DATA_BLOCK "DB_Z256_Scada"   // DB2010
{ S7_Optimized_Access := 'FALSE' }
VERSION : 0.1
   VAR
      tAlm : Struct   // HMI Alarms
         tE : Struct
            x0 : Bool;   // KE.Main emergency on
            x1 : Bool;   // KE1.Local emergency on
            x2 : Bool;   // Cabinet.Emergency localization
            x3 : Bool;   // SB1.Emergency localization
            x4 : Bool;   // SB2.Emergency localization
            x5 : Bool;
            x6 : Bool;
            x7 : Bool;
            x8 : Bool;
            x9 : Bool;
            x10 : Bool;
            x11 : Bool;
            x12 : Bool;
            x13 : Bool;
            x14 : Bool;
            x15 : Bool;
            x16 : Bool;
            x17 : Bool;
            x18 : Bool;
            x19 : Bool;
            x20 : Bool;
            x21 : Bool;
            x22 : Bool;
            x23 : Bool;
            x24 : Bool;
            x25 : Bool;
            x26 : Bool;
            x27 : Bool;
            x28 : Bool;
            x29 : Bool;
            x30 : Bool;
            x31 : Bool;
         END_STRUCT;
         tS : Struct
            tS0 : Struct
               x0 : Bool;   // xB18-3L+.PowerSupplyInputControlCabinetON
               x1 : Bool;   // xB18-7L+.InputInstallationPowerSupplyON"
               x2 : Bool;   // xB11QF1/1D/QF2.Anomaly power supplies 120V
               x3 : Bool;   // xB115KM1/2.AuxiliaryPowerSupplySetIn / xB18QF2.Power supply 24V logic
               x4 : Bool;   // xB410AP1.SafetyOnPanel1" / xB18QF3.Power supply 24V logic
               x5 : Bool;   // xB410AP1.SafetyOnPanel2" / xB20QF2.Power supply 24V logic
               x6 : Bool;   // xB20QF3.Power supply 24V logic
               x7 : Bool;   // xB21QF1.Power supply 24V logic
               x8 : Bool;   // xB140QF2.ProtectionPowerSupplyMotorsYcut" / xB41QF1.ProtectionPowerSupplyMotorsYcut 1-4
               x9 : Bool;   // xB41QF2.Protection power supply motors longitudinal cutting / xB41QF2.Protection power supply 36V motors longitudinal cutting 1-4
               x10 : Bool;   // xB42QF1.Protection power supply 36V / xB42QF1.ProtectionPowerSupplyMotorsYcut 5-8
               x11 : Bool;   // xB42QF2.Protection power supply motors longitudinal cutting / xB42QF2.Protection power supply 36V motors longitudinal cutting 5-8
               x12 : Bool;
               x13 : Bool;
               x14 : Bool;
               x15 : Bool;
               x16 : Bool;   // PLCA.Timeout receiving consumed message
               x17 : Bool;   // PLCB.Timeout receiving consumed message
               x18 : Bool;   // PLCA.Mission packet lost
               x19 : Bool;   // PLCB.Mission packet lost
               x20 : Bool;   // PLCA.Syncro packet lost
               x21 : Bool;   // PLCB.Syncro packet lost
               x22 : Bool;   // Syncro.YCut meter gap outside the limits
               x23 : Bool;   // Syncro.Main line meter gap outside the limits
               x24 : Bool;   // Syncro.Timeout receiving meter signal from main line
               x25 : Bool;   // Syncro.Timeout receiving syncro value from mainline
               x26 : Bool;   // Syncro.Unexpected syncro pulse
               x27 : Bool;   // Syncro.Unexpected syncro message
               x28 : Bool;   // Syncro.Machine not syncronized
               x29 : Bool;
               x30 : Bool;
               x31 : Bool;
            END_STRUCT;
            tS1 : Struct
               x0 : Bool;
               x1 : Bool;   // Syncro.YCut meter gap outside the limits
               x2 : Bool;
               x3 : Bool;
               x4 : Bool;
               x5 : Bool;
               x6 : Bool;
               x7 : Bool;
               x8 : Bool;   // xB21QF1.Power supply 24V logic
               x9 : Bool;
               x10 : Bool;   // Syncro.Main line meter gap outside the limits
               x11 : Bool;
               x12 : Bool;
               x13 : Bool;
               x14 : Bool;
               x15 : Bool;
               x16 : Bool;
               x17 : Bool;
               x18 : Bool;
               x19 : Bool;
               x20 : Bool;
               x21 : Bool;
               x22 : Bool;
               x23 : Bool;
               x24 : Bool;
               x25 : Bool;
               x26 : Bool;
               x27 : Bool;
               x28 : Bool;
               x29 : Bool;
               x30 : Bool;
               x31 : Bool;
            END_STRUCT;
            tS2 : Struct
               x0 : Bool;
               x1 : Bool;   // Syncro.YCut meter gap outside the limits
               x2 : Bool;
               x3 : Bool;
               x4 : Bool;
               x5 : Bool;
               x6 : Bool;
               x7 : Bool;
               x8 : Bool;   // xB21QF1.Power supply 24V logic
               x9 : Bool;
               x10 : Bool;   // Syncro.Main line meter gap outside the limits
               x11 : Bool;
               x12 : Bool;
               x13 : Bool;
               x14 : Bool;
               x15 : Bool;
               x16 : Bool;
               x17 : Bool;
               x18 : Bool;
               x19 : Bool;
               x20 : Bool;
               x21 : Bool;
               x22 : Bool;
               x23 : Bool;
               x24 : Bool;
               x25 : Bool;
               x26 : Bool;
               x27 : Bool;
               x28 : Bool;
               x29 : Bool;
               x30 : Bool;
               x31 : Bool;
            END_STRUCT;
            tS3 : Struct
               x0 : Bool;
               x1 : Bool;   // Syncro.YCut meter gap outside the limits
               x2 : Bool;
               x3 : Bool;
               x4 : Bool;
               x5 : Bool;
               x6 : Bool;
               x7 : Bool;
               x8 : Bool;   // xB21QF1.Power supply 24V logic
               x9 : Bool;
               x10 : Bool;   // Syncro.Main line meter gap outside the limits
               x11 : Bool;
               x12 : Bool;
               x13 : Bool;
               x14 : Bool;
               x15 : Bool;
               x16 : Bool;
               x17 : Bool;
               x18 : Bool;
               x19 : Bool;
               x20 : Bool;
               x21 : Bool;
               x22 : Bool;
               x23 : Bool;
               x24 : Bool;
               x25 : Bool;
               x26 : Bool;
               x27 : Bool;
               x28 : Bool;
               x29 : Bool;
               x30 : Bool;
               x31 : Bool;
            END_STRUCT;
         END_STRUCT;
         tF : Struct
            x0 : Bool;
            x1 : Bool;
            x2 : Bool;
            x3 : Bool;
            x4 : Bool;
            x5 : Bool;
            x6 : Bool;
            x7 : Bool;
            x8 : Bool;
            x9 : Bool;
            x10 : Bool;
            x11 : Bool;
            x12 : Bool;
            x13 : Bool;
            x14 : Bool;
            x15 : Bool;
            x16 : Bool;
            x17 : Bool;
            x18 : Bool;
            x19 : Bool;
            x20 : Bool;
            x21 : Bool;
            x22 : Bool;
            x23 : Bool;
            x24 : Bool;
            x25 : Bool;
            x26 : Bool;
            x27 : Bool;
            x28 : Bool;
            x29 : Bool;
            x30 : Bool;
            x31 : Bool;
         END_STRUCT;
         tW : Struct
            x0 : Bool;   // PLCA.Timeout receiving consumed message
            x1 : Bool;   // PLCB.Timeout receiving consumed message
            x2 : Bool;   // PLCA.Mission packet lost
            x3 : Bool;   // PLCB.Mission packet lost
            x4 : Bool;   // PLCA.Syncro packet lost
            x5 : Bool;   // PLCB.Syncro packet lost
            x6 : Bool;   // QF.Protection air conditioners
            x7 : Bool;
            x8 : Bool;
            x9 : Bool;
            x10 : Bool;
            x11 : Bool;
            x12 : Bool;
            x13 : Bool;
            x14 : Bool;
            x15 : Bool;
            x16 : Bool;
            x17 : Bool;
            x18 : Bool;
            x19 : Bool;
            x20 : Bool;
            x21 : Bool;
            x22 : Bool;
            x23 : Bool;
            x24 : Bool;
            x25 : Bool;
            x26 : Bool;
            x27 : Bool;
            x28 : Bool;
            x29 : Bool;
            x30 : Bool;
            x31 : Bool;
         END_STRUCT;
      END_STRUCT;
      tHMR : Struct   // HMI Read
         xCalibrationsAllowed : Bool := FALSE;   // Calibration function allowed {x|x|x|x|O}
         xSpare1 : Bool;
         xSpare2 : Bool;
         xSpare3 : Bool;
         xSpare4 : Bool;
         xSpare5 : Bool;
         xSpare6 : Bool;
         xSpare7 : Bool;
         xSpare8 : Bool;
         xSpare9 : Bool;
         xSpare10 : Bool;
         xSpare11 : Bool;
         xSpare12 : Bool;
         xSpare13 : Bool;
         xSpare14 : Bool;
         xZoneAlarm : Bool := FALSE;   // Zone alarm {X|X|X|X|O}
         xSpare16 : Bool;
         xSpare17 : Bool;
         xSpare18 : Bool;
         xSpare19 : Bool;
         xSpare20 : Bool;
         xSpare21 : Bool;
         xSpare22 : Bool;
         xSpare23 : Bool;
         xSpare24 : Bool;
         xSpare25 : Bool;
         xSpare26 : Bool;
         xSpare27 : Bool;
         xSpare28 : Bool;
         xSpare29 : Bool;
         xSpare30 : Bool;
         xSpare31 : Bool;
         xSpare : Array[0..15] of Bool;
         iSpare0 : Int;
         iSpare1 : Int;
         iSpare2 : Int;
         iSpare3 : Int;
         iSpare4 : Int;
         iSpare5 : Int;
         iSpare6 : Int;
         iSpare7 : Int;
         iSpare8 : Int;
         iSpare9 : Int;
         iSpare10 : Int;
         iSpare11 : Int;
         iSpare12 : Int;
         iSpare13 : Int;
         iSpare14 : Int;
         iSpare15 : Int;
         iSpare16 : Int;
         dZoneMode : DInt := 4;   // Zone modality (1=Manual;4=Automatic;8=Manual request) {x|x|x|x|O}
         dZoneState : DInt := 1024;   // Zone status (1=CycleON 2=StopCyc 4=CycleReq 8=StopReq 1024=E-Stop) {X|X|X|X|O} / HMI Alarms
         dCabinetStatusMCC : DInt := 1;   // Cabinet status MCC1256B (1=OK;2=General power alarm;3=Local power alarm) {X|X|X|X|O} / HMI Write
         dProdModeRequest : DInt := 3;   // Production modality request (1=Out of Production 3= In production) {x|x|x|x|O}
         dProdModeActual : DInt := 3;   // Production modality actual (1=Out of production 3=In production 8=Out of production request 9=In production request) {x|x|x|x|O}
         dSpare5 : DInt;
         "rgdHeadsActualStatus[0]" : DInt := 3;   // Head #1 prod. status (1=Out of production 3=In production 8=Out of production request 9=In production request) {x|x|x|x|O}
         "rgdHeadsActualStatus[1]" : DInt := 3;   // Head #2 prod. status (1=Out of production 3=In production 8=Out of production request 9=In production request) {x|x|x|x|O}
         "rgdHeadsActualStatus[2]" : DInt := 3;   // Head #3 prod. status (1=Out of production 3=In production 8=Out of production request 9=In production request) {x|x|x|x|O}
         "rgdHeadsActualStatus[3]" : DInt := 3;   // Head #4 prod. status (1=Out of production 3=In production 8=Out of production request 9=In production request) {x|x|x|x|O}
         "rgdHeadsActualStatus[4]" : DInt;   // Head #5 prod. status (1=Out of production 3=In production 8=Out of production request 9=In production request) {x|x|x|x|O}
         "rgdHeadsActualStatus[5]" : DInt;   // Head #6 prod. status (1=Out of production 3=In production 8=Out of production request 9=In production request) {x|x|x|x|O}
         "rgdHeadsActualStatus[6]" : DInt;   // Head #7 prod. status (1=Out of production 3=In production 8=Out of production request 9=In production request) {x|x|x|x|O}
         "rgdHeadsActualStatus[7]" : DInt;   // Head #8 prod. status (1=Out of production 3=In production 8=Out of production request 9=In production request) {x|x|x|x|O}
         dSpare14 : DInt;
         dSpare15 : DInt;
         dSpare : Array[0..15] of DInt;
         rSpare0 : Real;
         rSpare1 : Real;
         rSpare2 : Real;
         rSpare3 : Real;
         rSpare4 : Real;
         rSpare5 : Real;
         rSpare6 : Real;
         rSpare7 : Real;
         rSpare8 : Real;
         tManCmd : Struct
            xSpare0 : Bool;
            xSpare1 : Bool;
            xSpare2 : Bool;
            xSpare3 : Bool;
            xSpare4 : Bool;
            xSpare5 : Bool;
            xSpare6 : Bool;
            xSpare7 : Bool;
            xSpare8 : Bool;
            xSpare9 : Bool;
            xSpare10 : Bool;
            xSpare11 : Bool;
            xSpare12 : Bool;
            xSpare13 : Bool;
            xSpare14 : Bool;
            xSpare15 : Bool;
            xSpare : Array[0..15] of Bool;
         END_STRUCT;
      END_STRUCT;
      tHMW : Struct   // HMI Write
         xAutoModeReq : Bool := FALSE;   // Automatic mode request {x|x|x|x|O}
         xManModeReq : Bool := FALSE;   // Manual mode request {x|x|x|x|O}
         xOutOfProdReq : Bool := FALSE;   // Bridge out of production request {x|x|x|x|O}
         xInProdReq : Bool := FALSE;   // Bridge in production request {x|x|x|x|O}
         xCutOnBreakEnabled : Bool := FALSE;   // Cut during glass break {x|x|x|x|O}
         xMotorsAndCardsInitialize : Bool := FALSE;   // Motors and cards initialize {x|x|x|x|M}
         xForceHeadsHoming : Bool := FALSE;   // Force the homing of the heads {x|x|x|x|M}
         xPositionCalibrationRequest : Bool := FALSE;   // Position calibration request {x|x|x|x|M}
         xBridgeOffsetCalibrationRequest : Bool := FALSE;   // Bridge offset calibration request {x|x|x|x|M}
         xSpare9 : Bool;
         xSpare10 : Bool;
         xSpare11 : Bool;
         xSpare12 : Bool;
         xSpare13 : Bool;
         xGeneralReset : Bool := FALSE;   // General reset {X|X|X|X|M}
         xFaultsReset : Bool := FALSE;   // Reset faults {X|X|X|X|O}
         xHeadEnabled_1 : Bool := TRUE;   // Head #1 enabled/disabled {x|x|x|x|O}
         xHeadEnabled_2 : Bool := TRUE;   // Head #2 enabled/disabled {x|x|x|x|O}
         xHeadEnabled_3 : Bool := TRUE;   // Head #3 enabled/disabled {x|x|x|x|O}
         xHeadEnabled_4 : Bool := TRUE;   // Head #4 enabled/disabled {x|x|x|x|O}
         xHeadEnabled_5 : Bool := TRUE;   // Head #5 enabled/disabled {x|x|x|x|O}
         xHeadEnabled_6 : Bool := TRUE;   // Head #6 enabled/disabled {x|x|x|x|O}
         xHeadEnabled_7 : Bool := TRUE;   // Head #7 enabled/disabled {x|x|x|x|O}
         xHeadEnabled_8 : Bool := TRUE;   // Head #8 enabled/disabled {x|x|x|x|O}
         xSpare24 : Bool;
         xSpare25 : Bool;
         xSpare26 : Bool;
         xSpare27 : Bool;
         xSpare28 : Bool;
         xSpare29 : Bool;
         xSpare30 : Bool;
         xSpare31 : Bool;
         xSpare : Array[0..15] of Bool;
         iSpare0 : Int;
         iSpare1 : Int;
         iSpare2 : Int;
         iSpare3 : Int;
         iSpare4 : Int;
         iSpare5 : Int;
         iSpare6 : Int;
         iSpare7 : Int;
         iSpare8 : Int;
         iSpare9 : Int;
         iSpare10 : Int;
         iSpare11 : Int;
         iSpare12 : Int;
         iSpare13 : Int;
         iSpare14 : Int;
         iSpare15 : Int;
         iSpare16 : Int;
         dNumberOfLites : DInt := 1;   // Calibration. number of lite on calibration {x|x|1|8|M}
         dMoveBridgeOffset_cmm : DInt := 0;   // Calibration. Move all the heads of this offset {mm/100|mm|-100|100|M}
         dPressureScalerOnSample_perc : DInt := 100;   // Pressure scaler during sample plate [%] {%|%|0|100|O}
         dSpare3 : DInt;
         dSpare4 : DInt;
         dSpare5 : DInt;
         dSpare6 : DInt;
         dSpare7 : DInt;
         dHead_Selected_1 : DInt;   // Calibration. head number selected Cut1 {x|x|1|11|M}
         dHead_Selected_2 : DInt;   // Calibration. head number selected Cut2 {x|x|1|11|M}
         dHead_Selected_3 : DInt;   // Calibration. head number selected Cut3{x|x|1|11|M}
         dHead_Selected_4 : DInt;   // Calibration. head number selected Cut4{x|x|1|11|M}
         dHead_Selected_5 : DInt;   // Calibration. head number selected Cut5{x|x|1|11|M}
         dHead_Selected_6 : DInt;   // Calibration. head number selected Cut6{x|x|1|11|M}
         dHead_Selected_7 : DInt;   // Calibration. head number selected Cut7{x|x|1|11|M}
         dHead_Selected_8 : DInt;   // Calibration. head number selected Cut8{x|x|1|11|M}
         dCutWidthTeo_cmm_1 : DInt;   // Calibration. cut width Lite 1 theorical [mm/100] {mm/100|mm|200|4000|M}
         dCutWidthTeo_cmm_2 : DInt;   // Calibration. cut width Lite 2 theorical [mm/100] {mm/100|mm|200|4000|M}
         dCutWidthTeo_cmm_3 : DInt;   // Calibration. cut width Lite 3 theorical [mm/100] {mm/100|mm|200|4000|M}
         dCutWidthTeo_cmm_4 : DInt;   // Calibration. cut width Lite 4 theorical [mm/100] {mm/100|mm|200|4000|M}
         dCutWidthTeo_cmm_5 : DInt;   // Calibration. cut width Lite 5 theorical [mm/100] {mm/100|mm|200|4000|M}
         dCutWidthTeo_cmm_6 : DInt;   // Calibration. cut width Lite 6 theorical [mm/100] {mm/100|mm|200|4000|M}
         dCutWidthTeo_cmm_7 : DInt;   // Calibration. cut width Lite 7 theorical [mm/100] {mm/100|mm|200|4000|M}
         dCutWidthTeo_cmm_8 : DInt;   // Calibration. cut width Lite 8 theorical [mm/100] {mm/100|mm|200|4000|M}
         dCutWidthReal_cmm_1 : DInt;   // Calibration. cut width Lite 1 real [mm/100] {mm/100|mm|200|4000|M}
         dCutWidthReal_cmm_2 : DInt;   // Calibration. cut width Lite 2 real [mm/100] {mm/100|mm|200|4000|M}
         dCutWidthReal_cmm_3 : DInt;   // Calibration. cut width Lite 3 real [mm/100] {mm/100|mm|200|4000|M}
         dCutWidthReal_cmm_4 : DInt;   // Calibration. cut width Lite 4 real [mm/100] {mm/100|mm|200|4000|M}
         dCutWidthReal_cmm_5 : DInt;   // Calibration. cut width Lite 5 real [mm/100] {mm/100|mm|200|4000|M}
         dCutWidthReal_cmm_6 : DInt;   // Calibration. cut width Lite 6 real [mm/100] {mm/100|mm|200|4000|M}
         dCutWidthReal_cmm_7 : DInt;   // Calibration. cut width Lite 7 real [mm/100] {mm/100|mm|200|4000|M}
         dCutWidthReal_cmm_8 : DInt;   // Calibration. cut width Lite 8 real [mm/100] {mm/100|mm|200|4000|M}
         dSpare32 : DInt;
         dSpare33 : DInt;
         dSpare34 : DInt;
         dSpare35 : DInt;
         dSpare36 : DInt;
         dSpare37 : DInt;
         dSpare38 : DInt;
         dSpare39 : DInt;
         dSpare : Array[0..19] of DInt;
         rSpare0 : Real;
         rSpare1 : Real;
         rSpare2 : Real;
         rSpare3 : Real;
         rSpare4 : Real;
         rSpare5 : Real;
         rSpare6 : Real;
         rSpare7 : Real;
         rSpare8 : Real;
         tManCmd : Struct
            xBrakeEngage : Bool := FALSE;   // Brake engage all heads {x|x|x|x|O}
            xBrakeRelease : Bool := FALSE;   // Brake release all heads {x|x|x|x|O}
            xSpare2 : Bool;
            xSpare3 : Bool;
            xSpare4 : Bool;
            xSpare5 : Bool;
            xSpare6 : Bool;
            xSpare7 : Bool;
            xSpare8 : Bool;
            xSpare9 : Bool;
            xSpare10 : Bool;
            xSpare11 : Bool;
            xSpare12 : Bool;
            xSpare13 : Bool;
            xSpare14 : Bool;
            xSpare15 : Bool;
            xSpare16 : Bool;
            xSpare17 : Bool;
            xSpare18 : Bool;
            xSpare19 : Bool;
            xSpare20 : Bool;
            xSpare21 : Bool;
            xSpare22 : Bool;
            xSpare23 : Bool;
            xSpare24 : Bool;
            xSpare25 : Bool;
            xSpare26 : Bool;
            xSpare27 : Bool;
            xSpare28 : Bool;
            xSpare29 : Bool;
            xSpare30 : Bool;
            xSpare31 : Bool;
         END_STRUCT;
      END_STRUCT;
   END_VAR
BEGIN
END_DATA_BLOCK

DATA_BLOCK "DB_M256M_Scada"   // DB2011
{ S7_Optimized_Access := 'FALSE' }
VERSION : 0.1
   VAR
      tAlm : Struct   // HMI Alarms
         tE : Struct
            x0 : Bool;   // KE.Main emergency on
            x1 : Bool;   // KE1.Local emergency on
            x2 : Bool;   // Cabinet.Emergency localization
            x3 : Bool;   // SB1.Emergency localization
            x4 : Bool;   // SB2.Emergency localization
            x5 : Bool;
            x6 : Bool;
            x7 : Bool;
            x8 : Bool;
            x9 : Bool;
            x10 : Bool;
            x11 : Bool;
            x12 : Bool;
            x13 : Bool;
            x14 : Bool;
            x15 : Bool;
            x16 : Bool;
            x17 : Bool;
            x18 : Bool;
            x19 : Bool;
            x20 : Bool;
            x21 : Bool;
            x22 : Bool;
            x23 : Bool;
            x24 : Bool;
            x25 : Bool;
            x26 : Bool;
            x27 : Bool;
            x28 : Bool;
            x29 : Bool;
            x30 : Bool;
            x31 : Bool;
         END_STRUCT;
         tS : Struct
            tS0 : Struct
               x0 : Bool;   // xB18-3L+.PowerSupplyInputControlCabinetON / Head#1.Initialization timeout
               x1 : Bool;   // xB140QF2.ProtectionPowerSupplyMotorsYcut" / Head#1.homing timeout
               x2 : Bool;   // PLCA.Timeout receiving consumed message / Head#1.positioning timeout
               x3 : Bool;   // Syncro.Timeout receiving meter signal from main line / Head#1.carriage overload
               x4 : Bool;   // Head#1.drive error
               x5 : Bool;   // Head#1.missing ethernet IP connection
               x6 : Bool;   // Head#1.op.side overstroke
               x7 : Bool;   // Head#1.oppo.op.side overstroke
               x8 : Bool;   // Head#1.overstroke
               x9 : Bool;   // xB18-7L+.InputInstallationPowerSupplyON" / Head#2.Initialization timeout
               x10 : Bool;   // xB41QF2.Protection power supply motors longitudinal cutting / Head#2.homing timeout
               x11 : Bool;   // PLCB.Timeout receiving consumed message / Head#2.positioning timeout
               x12 : Bool;   // Syncro.Timeout receiving syncro value from mainline / Head#2.carriage overload
               x13 : Bool;   // Head#2.drive error
               x14 : Bool;   // Head#2.missing ethernet IP connection
               x15 : Bool;   // Head#2.op.side overstroke
               x16 : Bool;   // Head#2.oppo.op.side overstroke
               x17 : Bool;   // Head#2.overstroke
               x18 : Bool;   // xB11QF1/1D/QF2.Anomaly power supplies 120V / Head#3.Initialization timeout
               x19 : Bool;   // PLCA.Mission packet lost / Head#3.homing timeout
               x20 : Bool;   // Syncro.Unexpected syncro pulse / Head#3.positioning timeout
               x21 : Bool;   // Head#3.carriage overload
               x22 : Bool;   // Head#3.drive error
               x23 : Bool;   // Head#3.missing ethernet IP connection
               x24 : Bool;   // Head#3.op.side overstroke
               x25 : Bool;   // Head#3.oppo.op.side overstroke
               x26 : Bool;   // xB115KM1/2.AuxiliaryPowerSupplySetIn / Head#3.overstroke
               x27 : Bool;
               x28 : Bool;
               x29 : Bool;
               x30 : Bool;
               x31 : Bool;
            END_STRUCT;
            tS1 : Struct
               x0 : Bool;   // xB42QF2.Protection power supply motors longitudinal cutting / Head#4.Initialization timeout
               x1 : Bool;   // PLCB.Mission packet lost / Head#4.homing timeout
               x2 : Bool;   // Syncro.Unexpected syncro message / Head#4.positioning timeout
               x3 : Bool;   // Head#4.carriage overload
               x4 : Bool;   // Head#4.drive error
               x5 : Bool;   // Head#4.missing ethernet IP connection
               x6 : Bool;   // Head#4.op.side overstroke
               x7 : Bool;   // Head#4.oppo.op.side overstroke
               x8 : Bool;   // xB410AP1.SafetyOnPanel1" / Head#4.overstroke
               x9 : Bool;   // Head#5.Initialization timeout
               x10 : Bool;   // PLCA.Syncro packet lost / Head#5.homing timeout
               x11 : Bool;   // Syncro.Machine not syncronized / Head#5.positioning timeout
               x12 : Bool;   // Head#5.carriage overload
               x13 : Bool;   // Head#5.drive error
               x14 : Bool;   // Head#5.missing ethernet IP connection
               x15 : Bool;   // Head#5.op.side overstroke
               x16 : Bool;   // Head#5.oppo.op.side overstroke
               x17 : Bool;   // xB410AP1.SafetyOnPanel2" / Head#5.overstroke
               x18 : Bool;   // Head#6.Initialization timeout
               x19 : Bool;   // PLCB.Syncro packet lost / Head#6.homing timeout
               x20 : Bool;   // Head#6.positioning timeout
               x21 : Bool;   // Head#6.carriage overload
               x22 : Bool;   // Head#6.drive error
               x23 : Bool;   // Head#6.missing ethernet IP connection
               x24 : Bool;   // Head#6.op.side overstroke
               x25 : Bool;   // Head#6.oppo.op.side overstroke
               x26 : Bool;   // xB20QF3.Power supply 24V logic / Head#6.overstroke
               x27 : Bool;
               x28 : Bool;
               x29 : Bool;
               x30 : Bool;
               x31 : Bool;
            END_STRUCT;
            tS2 : Struct
               x0 : Bool;   // Head#7.Initialization timeout
               x1 : Bool;   // Syncro.YCut meter gap outside the limits / Head#7.homing timeout
               x2 : Bool;   // Head#7.positioning timeout
               x3 : Bool;   // Head#7.carriage overload
               x4 : Bool;   // Head#7.drive error
               x5 : Bool;   // Head#7.missing ethernet IP connection
               x6 : Bool;   // Head#7.op.side overstroke
               x7 : Bool;   // Head#7.oppo.op.side overstroke
               x8 : Bool;   // xB21QF1.Power supply 24V logic / Head#7.overstroke
               x9 : Bool;   // Head#8.Initialization timeout
               x10 : Bool;   // Syncro.Main line meter gap outside the limits / Head#8.homing timeout
               x11 : Bool;   // Head#8.positioning timeout
               x12 : Bool;   // Head#8.carriage overload
               x13 : Bool;   // Head#8.drive error
               x14 : Bool;   // Head#8.missing ethernet IP connection
               x15 : Bool;   // Head#8.op.side overstroke
               x16 : Bool;   // Head#8.oppo.op.side overstroke
               x17 : Bool;   // Head#8.overstroke
               x18 : Bool;
               x19 : Bool;
               x20 : Bool;
               x21 : Bool;
               x22 : Bool;
               x23 : Bool;
               x24 : Bool;
               x25 : Bool;
               x26 : Bool;
               x27 : Bool;
               x28 : Bool;
               x29 : Bool;
               x30 : Bool;
               x31 : Bool;
            END_STRUCT;
            tS3 : Struct
               x0 : Bool;
               x1 : Bool;   // Syncro.YCut meter gap outside the limits
               x2 : Bool;
               x3 : Bool;
               x4 : Bool;
               x5 : Bool;
               x6 : Bool;
               x7 : Bool;
               x8 : Bool;   // xB21QF1.Power supply 24V logic
               x9 : Bool;
               x10 : Bool;   // Syncro.Main line meter gap outside the limits
               x11 : Bool;
               x12 : Bool;
               x13 : Bool;
               x14 : Bool;
               x15 : Bool;
               x16 : Bool;
               x17 : Bool;
               x18 : Bool;
               x19 : Bool;
               x20 : Bool;
               x21 : Bool;
               x22 : Bool;
               x23 : Bool;
               x24 : Bool;
               x25 : Bool;
               x26 : Bool;
               x27 : Bool;
               x28 : Bool;
               x29 : Bool;
               x30 : Bool;
               x31 : Bool;
            END_STRUCT;
         END_STRUCT;
         tF : Struct
            x0 : Bool;
            x1 : Bool;
            x2 : Bool;
            x3 : Bool;
            x4 : Bool;
            x5 : Bool;
            x6 : Bool;
            x7 : Bool;
            x8 : Bool;
            x9 : Bool;
            x10 : Bool;
            x11 : Bool;
            x12 : Bool;
            x13 : Bool;
            x14 : Bool;
            x15 : Bool;
            x16 : Bool;
            x17 : Bool;
            x18 : Bool;
            x19 : Bool;
            x20 : Bool;
            x21 : Bool;
            x22 : Bool;
            x23 : Bool;
            x24 : Bool;
            x25 : Bool;
            x26 : Bool;
            x27 : Bool;
            x28 : Bool;
            x29 : Bool;
            x30 : Bool;
            x31 : Bool;
         END_STRUCT;
         tW : Struct
            x0 : Bool;   // PLCA.Timeout receiving consumed message
            x1 : Bool;   // PLCB.Timeout receiving consumed message
            x2 : Bool;   // PLCA.Mission packet lost
            x3 : Bool;   // PLCB.Mission packet lost
            x4 : Bool;   // PLCA.Syncro packet lost
            x5 : Bool;   // PLCB.Syncro packet lost
            x6 : Bool;   // QF.Protection air conditioners
            x7 : Bool;
            x8 : Bool;
            x9 : Bool;
            x10 : Bool;
            x11 : Bool;
            x12 : Bool;
            x13 : Bool;
            x14 : Bool;
            x15 : Bool;
            x16 : Bool;
            x17 : Bool;
            x18 : Bool;
            x19 : Bool;
            x20 : Bool;
            x21 : Bool;
            x22 : Bool;
            x23 : Bool;
            x24 : Bool;
            x25 : Bool;
            x26 : Bool;
            x27 : Bool;
            x28 : Bool;
            x29 : Bool;
            x30 : Bool;
            x31 : Bool;
         END_STRUCT;
      END_STRUCT;
      tHMR : Struct   // HMI Read
         xSpare0 : Bool := FALSE;   // Calibration function allowed {x|x|x|x|O}
         xSpare1 : Bool;
         xSpare2 : Bool;
         xSpare3 : Bool;
         xSpare4 : Bool;
         xSpare5 : Bool;
         xSpare6 : Bool;
         xSpare7 : Bool;
         xSpare8 : Bool;
         xSpare9 : Bool;
         xSpare10 : Bool;
         xSpare11 : Bool;
         xSpare12 : Bool;
         xSpare13 : Bool;
         xSpare14 : Bool;
         xSpare15 : Bool := FALSE;
         xSpare16 : Bool;
         xSpare17 : Bool;
         xSpare18 : Bool;
         xSpare19 : Bool;
         xSpare20 : Bool;
         xSpare21 : Bool;
         xSpare22 : Bool;
         xSpare23 : Bool;
         xSpare24 : Bool;
         xSpare25 : Bool;
         xSpare26 : Bool;
         xSpare27 : Bool;
         xSpare28 : Bool;
         xSpare29 : Bool;
         xSpare30 : Bool;
         xSpare31 : Bool;
         xSpare : Array[0..15] of Bool;
         iCodeAlarm_H1 : Int;   // Motor error code H1
         iCodeAlarm_H2 : Int;   // Motor error code H2
         iCodeAlarm_H3 : Int;   // Motor error code H3
         iCodeAlarm_H4 : Int;   // Motor error code H4
         iCodeAlarm_H5 : Int;   // Motor error code H5
         iCodeAlarm_H6 : Int;   // Motor error code H6
         iCodeAlarm_H7 : Int;   // Motor error code H7
         iCodeAlarm_H8 : Int;   // Motor error code H8
         iSpare8 : Int;
         iSpare9 : Int;
         iSpare10 : Int;
         iSpare11 : Int;
         iSpare12 : Int;
         iSpare13 : Int;
         iSpare14 : Int;
         iSpare15 : Int;
         iSpare16 : Int;
         dHeadActualPositions_cmm_H1 : DInt;   // Head#x head actual position [mm/100] {mm/100|mm|x|x|O} / Head#1 head actual position [mm/100] {mm/100|mm|x|x|O}
         dHeadActualPositions_cmm_H2 : DInt;   // Head#x head actual position [mm/100] {mm/100|mm|x|x|O} / Head#2 head actual position [mm/100] {mm/100|mm|x|x|O}
         dHeadActualPositions_cmm_H3 : DInt;   // Head#x head actual position [mm/100] {mm/100|mm|x|x|O} / Head#3 head actual position [mm/100] {mm/100|mm|x|x|O}
         dHeadActualPositions_cmm_H4 : DInt;   // Head#x head actual position [mm/100] {mm/100|mm|x|x|O} / Head#4 head actual position [mm/100] {mm/100|mm|x|x|O}
         dHeadActualPositions_cmm_H5 : DInt;   // Head#x head actual position [mm/100] {mm/100|mm|x|x|O} / Head#5 head actual position [mm/100] {mm/100|mm|x|x|O}
         dHeadActualPositions_cmm_H6 : DInt;   // Head#x head actual position [mm/100] {mm/100|mm|x|x|O} / Head#6 head actual position [mm/100] {mm/100|mm|x|x|O}
         dHeadActualPositions_cmm_H7 : DInt;   // Head#x head actual position [mm/100] {mm/100|mm|x|x|O} / Head#7 head actual position [mm/100] {mm/100|mm|x|x|O}
         dHeadActualPositions_cmm_H8 : DInt;   // Head#x head actual position [mm/100] {mm/100|mm|x|x|O} / Head#8 head actual position [mm/100] {mm/100|mm|x|x|O}
         dHeadHomePositions_cmm_H1 : DInt;   // Head#x home position [mm/100] {mm/100|mm|x|x|O} / Head#1 home position [mm/100] {mm/100|mm|x|x|O}
         dHeadHomePositions_cmm_H2 : DInt;   // Head#x home position [mm/100] {mm/100|mm|x|x|O} / Head#2 home position [mm/100] {mm/100|mm|x|x|O}
         dHeadHomePositions_cmm_H3 : DInt;   // Head#x home position [mm/100] {mm/100|mm|x|x|O} / Head#3 home position [mm/100] {mm/100|mm|x|x|O}
         dHeadHomePositions_cmm_H4 : DInt;   // Head#x home position [mm/100] {mm/100|mm|x|x|O} / Head#4 home position [mm/100] {mm/100|mm|x|x|O}
         dHeadHomePositions_cmm_H5 : DInt;   // Head#x home position [mm/100] {mm/100|mm|x|x|O} / Head#5 home position [mm/100] {mm/100|mm|x|x|O}
         dHeadHomePositions_cmm_H6 : DInt;   // Head#x home position [mm/100] {mm/100|mm|x|x|O} / Head#6 home position [mm/100] {mm/100|mm|x|x|O}
         dHeadHomePositions_cmm_H7 : DInt;   // Head#x home position [mm/100] {mm/100|mm|x|x|O} / Head#7 home position [mm/100] {mm/100|mm|x|x|O}
         dHeadHomePositions_cmm_H8 : DInt;   // Head#x home position [mm/100] {mm/100|mm|x|x|O} / Head#8 home position [mm/100] {mm/100|mm|x|x|O}
         dHeadMoveStatus_H1 : DInt;   // Head#x move status (1=Not Initialized 2=Not referred 3=Not positioned 4=Positioned 5=Positioning 6=Virtual collision 7=Anomaly) {x|x|x|x|O} / Head#1 move status (1=Not Initialized 2=Not referred 3=Not positioned 4=Positioned 5=Positioning 6=Virtual collision 7=Anomaly) {x|x|x|x|O}
         dHeadMoveStatus_H2 : DInt;   // Head#x move status (1=Not Initialized 2=Not referred 3=Not positioned 4=Positioned 5=Positioning 6=Virtual collision 7=Anomaly) {x|x|x|x|O} / Head#2 move status (1=Not Initialized 2=Not referred 3=Not positioned 4=Positioned 5=Positioning 6=Virtual collision 7=Anomaly) {x|x|x|x|O}
         dHeadMoveStatus_H3 : DInt;   // Head#x move status (1=Not Initialized 2=Not referred 3=Not positioned 4=Positioned 5=Positioning 6=Virtual collision 7=Anomaly) {x|x|x|x|O} / Head#3 move status (1=Not Initialized 2=Not referred 3=Not positioned 4=Positioned 5=Positioning 6=Virtual collision 7=Anomaly) {x|x|x|x|O}
         dHeadMoveStatus_H4 : DInt;   // Head#x move status (1=Not Initialized 2=Not referred 3=Not positioned 4=Positioned 5=Positioning 6=Virtual collision 7=Anomaly) {x|x|x|x|O} / Head#4 move status (1=Not Initialized 2=Not referred 3=Not positioned 4=Positioned 5=Positioning 6=Virtual collision 7=Anomaly) {x|x|x|x|O}
         dHeadMoveStatus_H5 : DInt;   // Head#x move status (1=Not Initialized 2=Not referred 3=Not positioned 4=Positioned 5=Positioning 6=Virtual collision 7=Anomaly) {x|x|x|x|O} / Head#5 move status (1=Not Initialized 2=Not referred 3=Not positioned 4=Positioned 5=Positioning 6=Virtual collision 7=Anomaly) {x|x|x|x|O}
         dHeadMoveStatus_H6 : DInt;   // Head#x move status (1=Not Initialized 2=Not referred 3=Not positioned 4=Positioned 5=Positioning 6=Virtual collision 7=Anomaly) {x|x|x|x|O} / Head#6 move status (1=Not Initialized 2=Not referred 3=Not positioned 4=Positioned 5=Positioning 6=Virtual collision 7=Anomaly) {x|x|x|x|O}
         dHeadMoveStatus_H7 : DInt;   // Head#x move status (1=Not Initialized 2=Not referred 3=Not positioned 4=Positioned 5=Positioning 6=Virtual collision 7=Anomaly) {x|x|x|x|O} / Head#7 move status (1=Not Initialized 2=Not referred 3=Not positioned 4=Positioned 5=Positioning 6=Virtual collision 7=Anomaly) {x|x|x|x|O}
         dHeadMoveStatus_H8 : DInt;   // Head#x move status (1=Not Initialized 2=Not referred 3=Not positioned 4=Positioned 5=Positioning 6=Virtual collision 7=Anomaly) {x|x|x|x|O} / Head#8 move status (1=Not Initialized 2=Not referred 3=Not positioned 4=Positioned 5=Positioning 6=Virtual collision 7=Anomaly) {x|x|x|x|O}
         dSpare : Array[0..7] of DInt;
         rSpare0 : Real;
         rSpare1 : Real;
         rSpare2 : Real;
         rSpare3 : Real;
         rSpare4 : Real;
         rSpare5 : Real;
         rSpare6 : Real;
         rSpare7 : Real;
         rSpare8 : Real;
         tManCmd : Struct
            xManJogForwardFdbk_H1 : Bool;   // Head#x manual jog forward fdbk {x|x|x|x|O} / Head#1 manual jog forward fdbk {x|x|x|x|O}
            xManJogBackwardFdbk_H1 : Bool;   // Head#x manual jog backward fdbk {x|x|x|x|O} / Head#1 manual jog backward fdbk {x|x|x|x|O}
            xManJogForwardFdbk_H2 : Bool;   // Head#x manual jog forward fdbk {x|x|x|x|O} / Head#2 manual jog forward fdbk {x|x|x|x|O}
            xManJogBackwardFdbk_H2 : Bool;   // Head#x manual jog backward fdbk {x|x|x|x|O} / Head#2 manual jog backward fdbk {x|x|x|x|O}
            xManJogForwardFdbk_H3 : Bool;   // Head#x manual jog forward fdbk {x|x|x|x|O} / Head#3 manual jog forward fdbk {x|x|x|x|O}
            xManJogBackwardFdbk_H3 : Bool;   // Head#x manual jog backward fdbk {x|x|x|x|O} / Head#3 manual jog backward fdbk {x|x|x|x|O}
            xManJogForwardFdbk_H4 : Bool;   // Head#x manual jog forward fdbk {x|x|x|x|O} / Head#4 manual jog forward fdbk {x|x|x|x|O}
            xManJogBackwardFdbk_H4 : Bool;   // Head#x manual jog backward fdbk {x|x|x|x|O} / Head#4 manual jog backward fdbk {x|x|x|x|O}
            xManJogForwardFdbk_H5 : Bool;   // Head#x manual jog forward fdbk {x|x|x|x|O} / Head#5 manual jog forward fdbk {x|x|x|x|O}
            xManJogBackwardFdbk_H5 : Bool;   // Head#x manual jog backward fdbk {x|x|x|x|O} / Head#5 manual jog backward fdbk {x|x|x|x|O}
            xManJogForwardFdbk_H6 : Bool;   // Head#x manual jog forward fdbk {x|x|x|x|O} / Head#6 manual jog forward fdbk {x|x|x|x|O}
            xManJogBackwardFdbk_H6 : Bool;   // Head#x manual jog backward fdbk {x|x|x|x|O} / Head#6 manual jog backward fdbk {x|x|x|x|O}
            xManJogForwardFdbk_H7 : Bool;   // Head#x manual jog forward fdbk {x|x|x|x|O} / Head#7 manual jog forward fdbk {x|x|x|x|O}
            xManJogBackwardFdbk_H7 : Bool;   // Head#x manual jog backward fdbk {x|x|x|x|O} / Head#7 manual jog backward fdbk {x|x|x|x|O}
            xManJogForwardFdbk_H8 : Bool;   // Head#x manual jog forward fdbk {x|x|x|x|O} / Head#8 manual jog forward fdbk {x|x|x|x|O}
            xManJogBackwardFdbk_H8 : Bool;   // Head#x manual jog backward fdbk {x|x|x|x|O} / Head#8 manual jog backward fdbk {x|x|x|x|O}
            xSpare : Array[0..15] of Bool;
         END_STRUCT;
      END_STRUCT;
      tHMW : Struct   // HMI Write
         xBrakeRealeaseHead_H1 : Bool := FALSE;   // Force the brake release of the head {x|x|x|x|M} / Force the brake release of the Head #1 {x|x|x|x|M}
         xBrakeEngageHeads_H1 : Bool := FALSE;   // Force the brake engaged of the head {x|x|x|x|M} / Force the brake engaged of the Head #1 {x|x|x|x|M}
         xUpdateHomeHead_H1 : Bool;   // Update home position head#x {x|x|x|x|M} / Update home position Head #1 {x|x|x|x|M}
         xBrakeRealeaseHead_H2 : Bool := FALSE;   // Force the brake release of the head {x|x|x|x|M} / Force the brake release of the Head #2 {x|x|x|x|M}
         xBrakeEngageHeads_H2 : Bool := FALSE;   // Force the brake engaged of the head {x|x|x|x|M} / Force the brake engaged of the Head #2 {x|x|x|x|M}
         xUpdateHomeHead_H2 : Bool;   // Update home position head#x {x|x|x|x|M} / Update home position Head #2 {x|x|x|x|M}
         xBrakeRealeaseHead_H3 : Bool := FALSE;   // Force the brake release of the head {x|x|x|x|M} / Force the brake release of the Head #3 {x|x|x|x|M}
         xBrakeEngageHeads_H3 : Bool := FALSE;   // Force the brake engaged of the head {x|x|x|x|M} / Force the brake engaged of the Head #3 {x|x|x|x|M}
         xUpdateHomeHead_H3 : Bool;   // Update home position head#x {x|x|x|x|M} / Update home position Head #3 {x|x|x|x|M}
         xBrakeRealeaseHead_H4 : Bool := FALSE;   // Force the brake release of the head {x|x|x|x|M} / Force the brake release of the Head #4{x|x|x|x|M}
         xBrakeEngageHeads_H4 : Bool := FALSE;   // Force the brake engaged of the head {x|x|x|x|M} / Force the brake engaged of the Head #4{x|x|x|x|M}
         xUpdateHomeHead_H4 : Bool;   // Update home position head#x {x|x|x|x|M} / Update home position Head #4 {x|x|x|x|M}
         xBrakeRealeaseHead_H5 : Bool := FALSE;   // Force the brake release of the head {x|x|x|x|M} / Force the brake release of the Head #5{x|x|x|x|M}
         xBrakeEngageHeads_H5 : Bool := FALSE;   // Force the brake engaged of the head {x|x|x|x|M} / Force the brake engaged of the Head #5{x|x|x|x|M}
         xUpdateHomeHead_H5 : Bool;   // Update home position head#x {x|x|x|x|M} / Update home position Head #5 {x|x|x|x|M}
         xBrakeRealeaseHead_H6 : Bool := FALSE;   // Force the brake release of the head {x|x|x|x|M} / Force the brake release of the Head #6{x|x|x|x|M}
         xBrakeEngageHeads_H6 : Bool := FALSE;   // Force the brake engaged of the head {x|x|x|x|M} / Force the brake engaged of the Head #6 {x|x|x|x|M}
         xUpdateHomeHead_H6 : Bool;   // Update home position head#x {x|x|x|x|M} / Update home position Head #6 {x|x|x|x|M}
         xBrakeRealeaseHead_H7 : Bool := FALSE;   // Force the brake release of the head {x|x|x|x|M} / Force the brake release of the Head #7{x|x|x|x|M}
         xBrakeEngageHeads_H7 : Bool := FALSE;   // Force the brake engaged of the head {x|x|x|x|M} / Force the brake engaged of the Head #7{x|x|x|x|M}
         xUpdateHomeHead_H7 : Bool;   // Update home position head#x {x|x|x|x|M} / Update home position Head #7{x|x|x|x|M}
         xBrakeRealeaseHead_H8 : Bool := FALSE;   // Force the brake release of the head {x|x|x|x|M} / Force the brake release of the Head #8{x|x|x|x|M}
         xBrakeEngageHeads_H8 : Bool := FALSE;   // Force the brake engaged of the head {x|x|x|x|M} / Force the brake engaged of the Head #8{x|x|x|x|M}
         xUpdateHomeHead_H8 : Bool;   // Update home position head#x {x|x|x|x|M} / Update home position Head #8 {x|x|x|x|M}
         xSpare24 : Bool;
         xSpare25 : Bool;
         xSpare26 : Bool;
         xSpare27 : Bool;
         xSpare28 : Bool;
         xSpare29 : Bool;
         xSpare30 : Bool;
         xSpare31 : Bool;
         xSpare : Array[0..15] of Bool;
         iSpare0 : Int;
         iSpare1 : Int;
         iSpare2 : Int;
         iSpare3 : Int;
         iSpare4 : Int;
         iSpare5 : Int;
         iSpare6 : Int;
         iSpare7 : Int;
         iSpare8 : Int;
         iSpare9 : Int;
         iSpare10 : Int;
         iSpare11 : Int;
         iSpare12 : Int;
         iSpare13 : Int;
         iSpare14 : Int;
         iSpare15 : Int;
         iSpare16 : Int;
         dHeadHomePositions_cmm_H1 : DInt;   // Head#x home position [mm/100] {mm/100|mm|-2500|2500|M} / Head#1 home position [mm/100] {mm/100|mm|-2500|2500|M}
         dHeadHomePositions_cmm_H2 : DInt;   // Head#x home position [mm/100] {mm/100|mm|-2500|2500|M} / Head#2 home position [mm/100] {mm/100|mm|-2500|2500|M}
         dHeadHomePositions_cmm_H3 : DInt;   // Head#x home position [mm/100] {mm/100|mm|-2500|2500|M} / Head#3 home position [mm/100] {mm/100|mm|-2500|2500|M}
         dHeadHomePositions_cmm_H4 : DInt;   // Head#x home position [mm/100] {mm/100|mm|-2500|2500|M} / Head#4 home position [mm/100] {mm/100|mm|-2500|2500|M}
         dHeadHomePositions_cmm_H5 : DInt;   // Head#x home position [mm/100] {mm/100|mm|-2500|2500|M} / Head#5 home position [mm/100] {mm/100|mm|-2500|2500|M}
         dHeadHomePositions_cmm_H6 : DInt;   // Head#x home position [mm/100] {mm/100|mm|-2500|2500|M} / Head#6 home position [mm/100] {mm/100|mm|-2500|2500|M}
         dHeadHomePositions_cmm_H7 : DInt;   // Head#x home position [mm/100] {mm/100|mm|-2500|2500|M} / Head#7 home position [mm/100] {mm/100|mm|-2500|2500|M}
         dHeadHomePositions_cmm_H8 : DInt;   // Head#x home position [mm/100] {mm/100|mm|-2500|2500|M} / Head#8 home position [mm/100] {mm/100|mm|-2500|2500|M}
         dSpare8 : DInt;
         dSpare9 : DInt;
         dSpare10 : DInt;
         dSpare11 : DInt;
         dSpare12 : DInt;
         dSpare13 : DInt;
         dSpare14 : DInt;
         dSpare15 : DInt;
         dSpare : Array[0..43] of DInt;
         rSpare0 : Real;
         rSpare1 : Real;
         rSpare2 : Real;
         rSpare3 : Real;
         rSpare4 : Real;
         rSpare5 : Real;
         rSpare6 : Real;
         rSpare7 : Real;
         rSpare8 : Real;
         tManCmd : Struct
            xMan_JogForward_H1 : Bool;   // Head #x manual jog forward {x|x|x|x|O} / Head #1 manual jog forward {x|x|x|x|O}
            xMan_JogBackward_H1 : Bool;   // Head #x manual jog backward {x|x|x|x|O} / Head #1 manual jog backward {x|x|x|x|O}
            xMan_JogForward_H2 : Bool;   // Head #x manual jog forward {x|x|x|x|O} / Head #2 manual jog forward {x|x|x|x|O}
            xMan_JogBackward_H2 : Bool;   // Head #x manual jog backward {x|x|x|x|O} / Head #2 manual jog backward {x|x|x|x|O}
            xMan_JogForward_H3 : Bool;   // Head #x manual jog forward {x|x|x|x|O} / Head #3 manual jog forward {x|x|x|x|O}
            xMan_JogBackward_H3 : Bool;   // Head #x manual jog backward {x|x|x|x|O} / Head #3 manual jog backward {x|x|x|x|O}
            xMan_JogForward_H4 : Bool;   // Head #x manual jog forward {x|x|x|x|O} / Head #4 manual jog forward {x|x|x|x|O}
            xMan_JogBackward_H4 : Bool;   // Head #x manual jog backward {x|x|x|x|O} / Head #4 manual jog backward {x|x|x|x|O}
            xMan_JogForward_H5 : Bool;   // Head #x manual jog forward {x|x|x|x|O} / Head #5 manual jog forward {x|x|x|x|O}
            xMan_JogBackward_H5 : Bool;   // Head #x manual jog backward {x|x|x|x|O} / Head #5 manual jog backward {x|x|x|x|O}
            xMan_JogForward_H6 : Bool;   // Head #x manual jog forward {x|x|x|x|O} / Head #6 manual jog forward {x|x|x|x|O}
            xMan_JogBackward_H6 : Bool;   // Head #x manual jog backward {x|x|x|x|O} / Head #6 manual jog backward {x|x|x|x|O}
            xMan_JogForward_H7 : Bool;   // Head #x manual jog forward {x|x|x|x|O} / Head #7 manual jog forward {x|x|x|x|O}
            xMan_JogBackward_H7 : Bool;   // Head #x manual jog backward {x|x|x|x|O} / Head #7 manual jog backward {x|x|x|x|O}
            xMan_JogForward_H8 : Bool;   // Head #x manual jog forward {x|x|x|x|O} / Head #8 manual jog forward {x|x|x|x|O}
            xMan_JogBackward_H8 : Bool;   // Head #x manual jog backward {x|x|x|x|O} / Head #8 manual jog backward {x|x|x|x|O}
            xSpare16 : Bool;
            xSpare17 : Bool;
            xSpare18 : Bool;
            xSpare19 : Bool;
            xSpare20 : Bool;
            xSpare21 : Bool;
            xSpare22 : Bool;
            xSpare23 : Bool;
            xSpare24 : Bool;
            xSpare25 : Bool;
            xSpare26 : Bool;
            xSpare27 : Bool;
            xSpare28 : Bool;
            xSpare29 : Bool;
            xSpare30 : Bool;
            xSpare31 : Bool;
         END_STRUCT;
      END_STRUCT;
   END_VAR
BEGIN
END_DATA_BLOCK

DATA_BLOCK "DB_M256F_Scada"   // DB2012
{ S7_Optimized_Access := 'FALSE' }